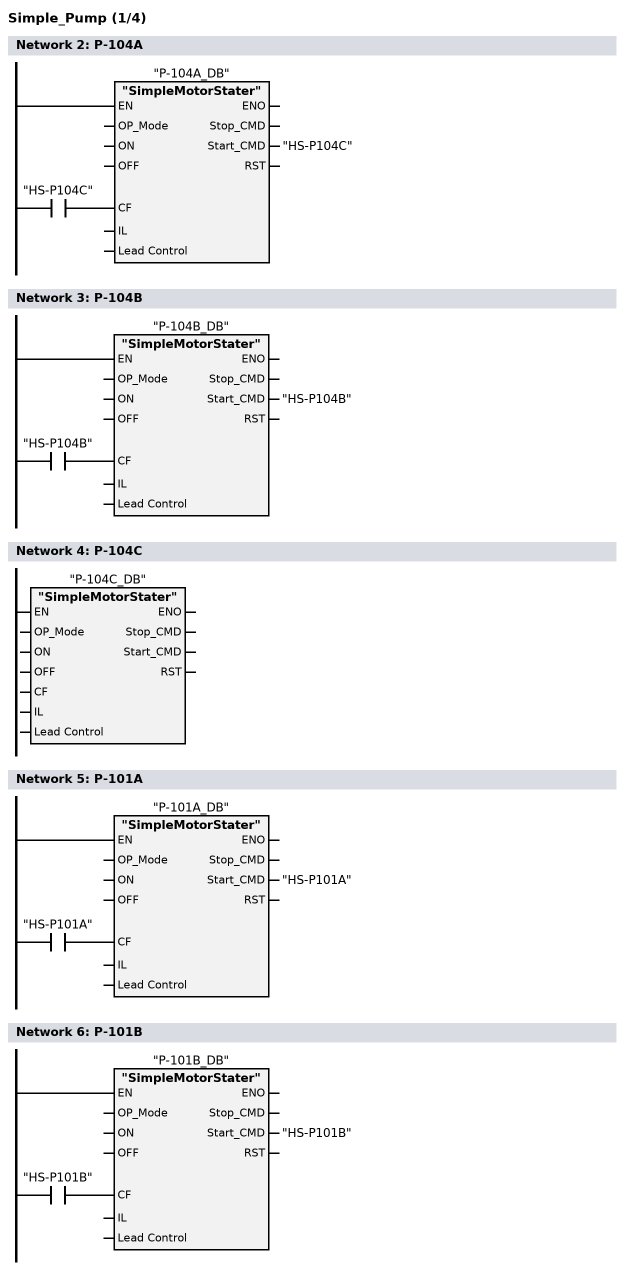
   RUNG wire#powerrail
      "P-104A_DB"(CF := wire#w1, OP_Mode :=, ON :=, OFF :=, IL :=, "Lead Control" :=, Stop_CMD =>, Start_CMD => "HS-P104C", RST =>)
   END_RUNG
   RUNG wire#powerrail
      Contact( "HS-P104C" )
   END_RUNG wire#w1
   // the same network as SCL:
   "P-104A_DB"(CF := "HS-P104C", Start_CMD => "HS-P104C");   // "SimpleMotorStater"
END_REGION

REGION Network 3: P-104B
   RUNG wire#powerrail
      "P-104B_DB"(CF := wire#w1, OP_Mode :=, ON :=, OFF :=, IL :=, "Lead Control" :=, Stop_CMD =>, Start_CMD => "HS-P104B", RST =>)
   END_RUNG
   RUNG wire#powerrail
      Contact( "HS-P104B" )
   END_RUNG wire#w1
   // the same network as SCL:
   "P-104B_DB"(CF := "HS-P104B", Start_CMD => "HS-P104B");   // "SimpleMotorStater"
END_REGION

REGION Network 4: P-104C
   RUNG wire#powerrail
      "P-104C_DB"(OP_Mode :=, ON :=, OFF :=, CF :=, IL :=, "Lead Control" :=, Stop_CMD =>, Start_CMD =>, RST =>)
   END_RUNG
   // the same network as SCL:
   "P-104C_DB"();   // "SimpleMotorStater"
END_REGION

REGION Network 5: P-101A
   RUNG wire#powerrail
      "P-101A_DB"(CF := wire#w1, OP_Mode :=, ON :=, OFF :=, IL :=, "Lead Control" :=, Stop_CMD =>, Start_CMD => "HS-P101A", RST =>)
   END_RUNG
   RUNG wire#powerrail
      Contact( "HS-P101A" )
   END_RUNG wire#w1
   // the same network as SCL:
   "P-101A_DB"(CF := "HS-P101A", Start_CMD => "HS-P101A");   // "SimpleMotorStater"
END_REGION

REGION Network 6: P-101B
   RUNG wire#powerrail
      "P-101B_DB"(CF := wire#w1, OP_Mode :=, ON :=, OFF :=, IL :=, "Lead Control" :=, Stop_CMD =>, Start_CMD => "HS-P101B", RST =>)
   END_RUNG
   RUNG wire#powerrail
      Contact( "HS-P101B" )
   END_RUNG wire#w1
   // the same network as SCL:
   "P-101B_DB"(CF := "HS-P101B", Start_CMD => "HS-P101B");   // "SimpleMotorStater"
END_REGION

REGION Network 7: P-102A
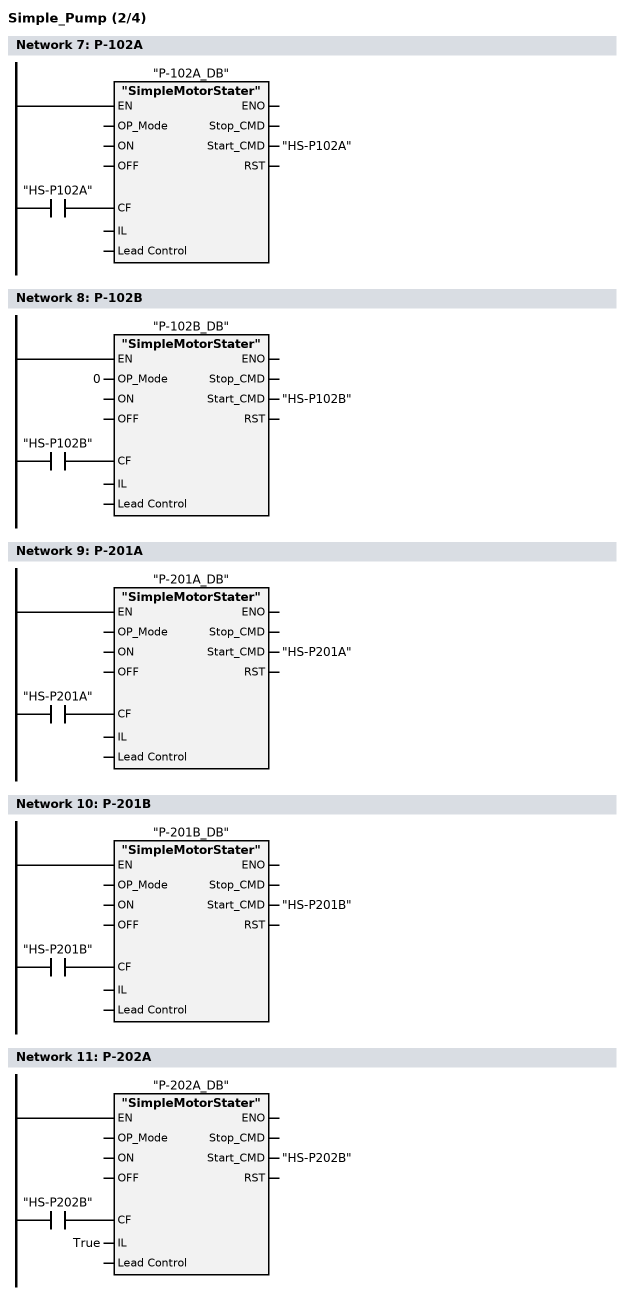
   RUNG wire#powerrail
      "P-102A_DB"(CF := wire#w1, OP_Mode :=, ON :=, OFF :=, IL :=, "Lead Control" :=, Stop_CMD =>, Start_CMD => "HS-P102A", RST =>)
   END_RUNG
   RUNG wire#powerrail
      Contact( "HS-P102A" )
   END_RUNG wire#w1
   // the same network as SCL:
   "P-102A_DB"(CF := "HS-P102A", Start_CMD => "HS-P102A");   // "SimpleMotorStater"
END_REGION

REGION Network 8: P-102B
   RUNG wire#powerrail
      "P-102B_DB"(CF := wire#w1, OP_Mode := 0, ON :=, OFF :=, IL :=, "Lead Control" :=, Stop_CMD =>, Start_CMD => "HS-P102B", RST =>)
   END_RUNG
   RUNG wire#powerrail
      Contact( "HS-P102B" )
   END_RUNG wire#w1
   // the same network as SCL:
   "P-102B_DB"(OP_Mode := 0, CF := "HS-P102B", Start_CMD => "HS-P102B");   // "SimpleMotorStater"
END_REGION

REGION Network 9: P-201A
   RUNG wire#powerrail
      "P-201A_DB"(CF := wire#w1, OP_Mode :=, ON :=, OFF :=, IL :=, "Lead Control" :=, Stop_CMD =>, Start_CMD => "HS-P201A", RST =>)
   END_RUNG
   RUNG wire#powerrail
      Contact( "HS-P201A" )
   END_RUNG wire#w1
   // the same network as SCL:
   "P-201A_DB"(CF := "HS-P201A", Start_CMD => "HS-P201A");   // "SimpleMotorStater"
END_REGION

REGION Network 10: P-201B
   RUNG wire#powerrail
      "P-201B_DB"(CF := wire#w1, OP_Mode :=, ON :=, OFF :=, IL :=, "Lead Control" :=, Stop_CMD =>, Start_CMD => "HS-P201B", RST =>)
   END_RUNG
   RUNG wire#powerrail
      Contact( "HS-P201B" )
   END_RUNG wire#w1
   // the same network as SCL:
   "P-201B_DB"(CF := "HS-P201B", Start_CMD => "HS-P201B");   // "SimpleMotorStater"
END_REGION

REGION Network 11: P-202A
   RUNG wire#powerrail
      "P-202A_DB"(CF := wire#w1, OP_Mode :=, ON :=, OFF :=, IL := True, "Lead Control" :=, Stop_CMD =>, Start_CMD => "HS-P202B", RST =>)
   END_RUNG
   RUNG wire#powerrail
      Contact( "HS-P202B" )
   END_RUNG wire#w1
   // the same network as SCL:
   "P-202A_DB"(CF := "HS-P202B", IL := True, Start_CMD => "HS-P202B");   // "SimpleMotorStater"
END_REGION

REGION Network 12: P-202B
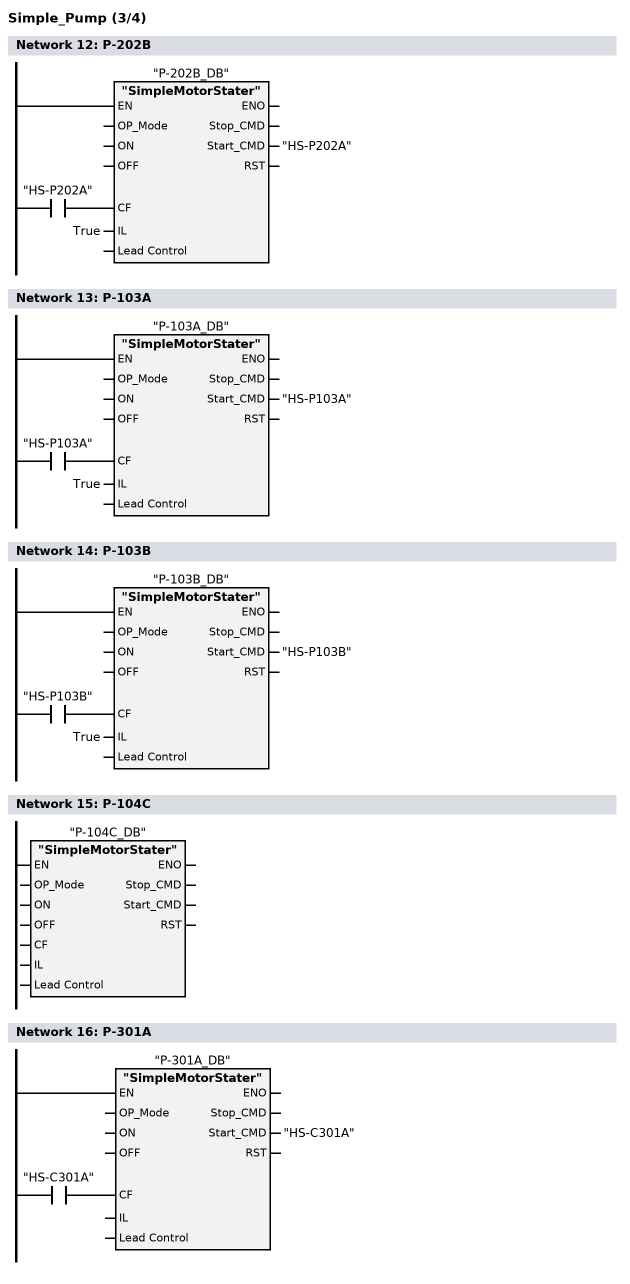
   RUNG wire#powerrail
      "P-202B_DB"(CF := wire#w1, OP_Mode :=, ON :=, OFF :=, IL := True, "Lead Control" :=, Stop_CMD =>, Start_CMD => "HS-P202A", RST =>)
   END_RUNG
   RUNG wire#powerrail
      Contact( "HS-P202A" )
   END_RUNG wire#w1
   // the same network as SCL:
   "P-202B_DB"(CF := "HS-P202A", IL := True, Start_CMD => "HS-P202A");   // "SimpleMotorStater"
END_REGION

REGION Network 13: P-103A
   RUNG wire#powerrail
      "P-103A_DB"(CF := wire#w1, OP_Mode :=, ON :=, OFF :=, IL := True, "Lead Control" :=, Stop_CMD =>, Start_CMD => "HS-P103A", RST =>)
   END_RUNG
   RUNG wire#powerrail
      Contact( "HS-P103A" )
   END_RUNG wire#w1
   // the same network as SCL:
   "P-103A_DB"(CF := "HS-P103A", IL := True, Start_CMD => "HS-P103A");   // "SimpleMotorStater"
END_REGION

REGION Network 14: P-103B
   RUNG wire#powerrail
      "P-103B_DB"(CF := wire#w1, OP_Mode :=, ON :=, OFF :=, IL := True, "Lead Control" :=, Stop_CMD =>, Start_CMD => "HS-P103B", RST =>)
   END_RUNG
   RUNG wire#powerrail
      Contact( "HS-P103B" )
   END_RUNG wire#w1
   // the same network as SCL:
   "P-103B_DB"(CF := "HS-P103B", IL := True, Start_CMD => "HS-P103B");   // "SimpleMotorStater"
END_REGION

REGION Network 15: P-104C
   RUNG wire#powerrail
      "P-104C_DB"(OP_Mode :=, ON :=, OFF :=, CF :=, IL :=, "Lead Control" :=, Stop_CMD =>, Start_CMD =>, RST =>)
   END_RUNG
   // the same network as SCL:
   "P-104C_DB"();   // "SimpleMotorStater"
END_REGION

REGION Network 16: P-301A
   RUNG wire#powerrail
      "P-301A_DB"(CF := wire#w1, OP_Mode :=, ON :=, OFF :=, IL :=, "Lead Control" :=, Stop_CMD =>, Start_CMD => "HS-C301A", RST =>)
   END_RUNG
   RUNG wire#powerrail
      Contact( "HS-C301A" )
   END_RUNG wire#w1
   // the same network as SCL:
   "P-301A_DB"(CF := "HS-C301A", Start_CMD => "HS-C301A");   // "SimpleMotorStater"
END_REGION

REGION Network 17: P-301B
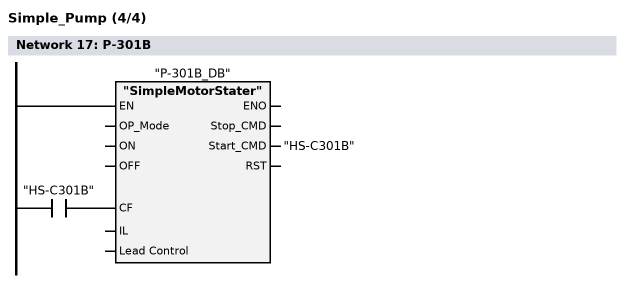
   RUNG wire#powerrail
      "P-301B_DB"(CF := wire#w1, OP_Mode :=, ON :=, OFF :=, IL :=, "Lead Control" :=, Stop_CMD =>, Start_CMD => "HS-C301B", RST =>)
   END_RUNG
   RUNG wire#powerrail
      Contact( "HS-C301B" )
   END_RUNG wire#w1
   // the same network as SCL:
   "P-301B_DB"(CF := "HS-C301B", Start_CMD => "HS-C301B");   // "SimpleMotorStater"
END_REGION
END_FUNCTION

// folder: Signal Digital Output/Centrifuge

FUNCTION "Centrifuge_DO" : Void   // FC108, LAD
{ S7_Optimized_Access := 'TRUE' }
VERSION : 0.1
BEGIN

REGION Network 1: Centrifuge Start Command
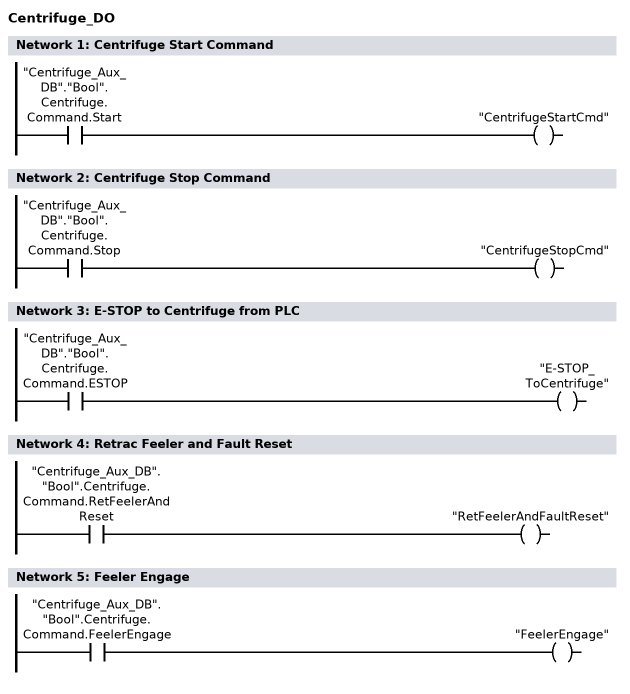
   RUNG wire#powerrail
      Contact( "Centrifuge_Aux_DB"."Bool".Centrifuge.Command.Start )
      Coil( "CentrifugeStartCmd" )
   END_RUNG
   // the same network as SCL:
   "CentrifugeStartCmd" := "Centrifuge_Aux_DB"."Bool".Centrifuge.Command.Start;
END_REGION

REGION Network 2: Centrifuge Stop Command
   RUNG wire#powerrail
      Contact( "Centrifuge_Aux_DB"."Bool".Centrifuge.Command.Stop )
      Coil( "CentrifugeStopCmd" )
   END_RUNG
   // the same network as SCL:
   "CentrifugeStopCmd" := "Centrifuge_Aux_DB"."Bool".Centrifuge.Command.Stop;
END_REGION

REGION Network 3: E-STOP to Centrifuge from PLC
   RUNG wire#powerrail
      Contact( "Centrifuge_Aux_DB"."Bool".Centrifuge.Command.ESTOP )
      Coil( "E-STOP_ToCentrifuge" )
   END_RUNG
   // the same network as SCL:
   "E-STOP_ToCentrifuge" := "Centrifuge_Aux_DB"."Bool".Centrifuge.Command.ESTOP;
END_REGION

REGION Network 4: Retrac Feeler and Fault Reset
   RUNG wire#powerrail
      Contact( "Centrifuge_Aux_DB"."Bool".Centrifuge.Command.RetFeelerAndReset )
      Coil( "RetFeelerAndFaultReset" )
   END_RUNG
   // the same network as SCL:
   "RetFeelerAndFaultReset" := "Centrifuge_Aux_DB"."Bool".Centrifuge.Command.RetFeelerAndReset;
END_REGION

REGION Network 5: Feeler Engage
   RUNG wire#powerrail
      Contact( "Centrifuge_Aux_DB"."Bool".Centrifuge.Command.FeelerEngage )
      Coil( "FeelerEngage" )
   END_RUNG
   // the same network as SCL:
   "FeelerEngage" := "Centrifuge_Aux_DB"."Bool".Centrifuge.Command.FeelerEngage;
END_REGION
END_FUNCTION

// folder: Signal Inputs

FUNCTION "Signals" : Void   // FC6, LAD
{ S7_Optimized_Access := 'TRUE' }
VERSION : 0.1
BEGIN

REGION Network 1: LSHH-1011 : T-101 High High Level Switch
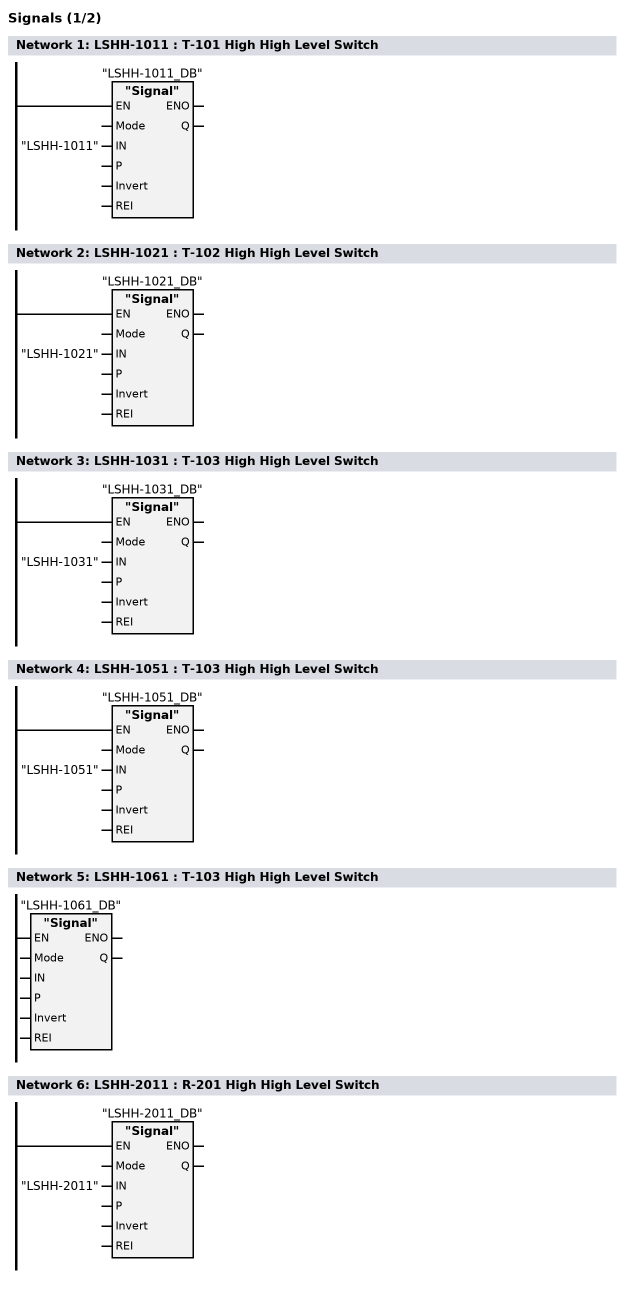
   RUNG wire#powerrail
      "LSHH-1011_DB"(Mode :=, IN := "LSHH-1011", P :=, Invert :=, REI :=, Q =>)
   END_RUNG
   // the same network as SCL:
   "LSHH-1011_DB"(IN := "LSHH-1011");   // "Signal"
END_REGION

REGION Network 2: LSHH-1021 : T-102 High High Level Switch
   RUNG wire#powerrail
      "LSHH-1021_DB"(Mode :=, IN := "LSHH-1021", P :=, Invert :=, REI :=, Q =>)
   END_RUNG
   // the same network as SCL:
   "LSHH-1021_DB"(IN := "LSHH-1021");   // "Signal"
END_REGION

REGION Network 3: LSHH-1031 : T-103 High High Level Switch
   RUNG wire#powerrail
      "LSHH-1031_DB"(Mode :=, IN := "LSHH-1031", P :=, Invert :=, REI :=, Q =>)
   END_RUNG
   // the same network as SCL:
   "LSHH-1031_DB"(IN := "LSHH-1031");   // "Signal"
END_REGION

REGION Network 4: LSHH-1051 : T-103 High High Level Switch
   RUNG wire#powerrail
      "LSHH-1051_DB"(Mode :=, IN := "LSHH-1051", P :=, Invert :=, REI :=, Q =>)
   END_RUNG
   // the same network as SCL:
   "LSHH-1051_DB"(IN := "LSHH-1051");   // "Signal"
END_REGION

REGION Network 5: LSHH-1061 : T-103 High High Level Switch
   RUNG wire#powerrail
      "LSHH-1061_DB"(Mode :=, IN :=, P :=, Invert :=, REI :=, Q =>)
   END_RUNG
   // the same network as SCL:
   "LSHH-1061_DB"();   // "Signal"
END_REGION

REGION Network 6: LSHH-2011 : R-201 High High Level Switch
   RUNG wire#powerrail
      "LSHH-2011_DB"(Mode :=, IN := "LSHH-2011", P :=, Invert :=, REI :=, Q =>)
   END_RUNG
   // the same network as SCL:
   "LSHH-2011_DB"(IN := "LSHH-2011");   // "Signal"
END_REGION

REGION Network 7: LSHH-2021 : R-202 High High Level Switch
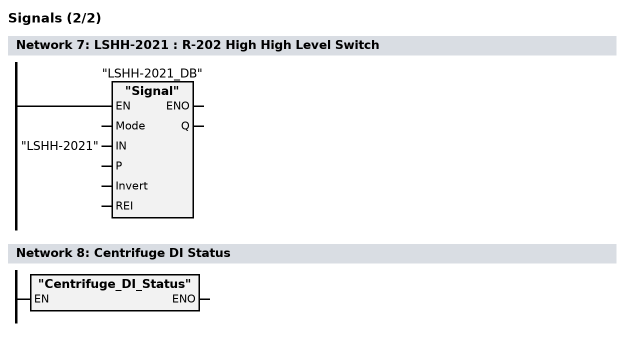
   RUNG wire#powerrail
      "LSHH-2021_DB"(Mode :=, IN := "LSHH-2021", P :=, Invert :=, REI :=, Q =>)
   END_RUNG
   // the same network as SCL:
   "LSHH-2021_DB"(IN := "LSHH-2021");   // "Signal"
END_REGION

REGION Network 8: Centrifuge DI Status
   RUNG wire#powerrail
      "Centrifuge_DI_Status"()
   END_RUNG
   // the same network as SCL:
   "Centrifuge_DI_Status"();
END_REGION
END_FUNCTION

// folder: Signal Inputs/Centrifuge

FUNCTION "Centrifuge_DI_Status" : Void   // FC104, LAD
{ S7_Optimized_Access := 'TRUE' }
VERSION : 0.1
// Digital Input from Centrifuge
BEGIN

REGION Network 1: Vibration Fault
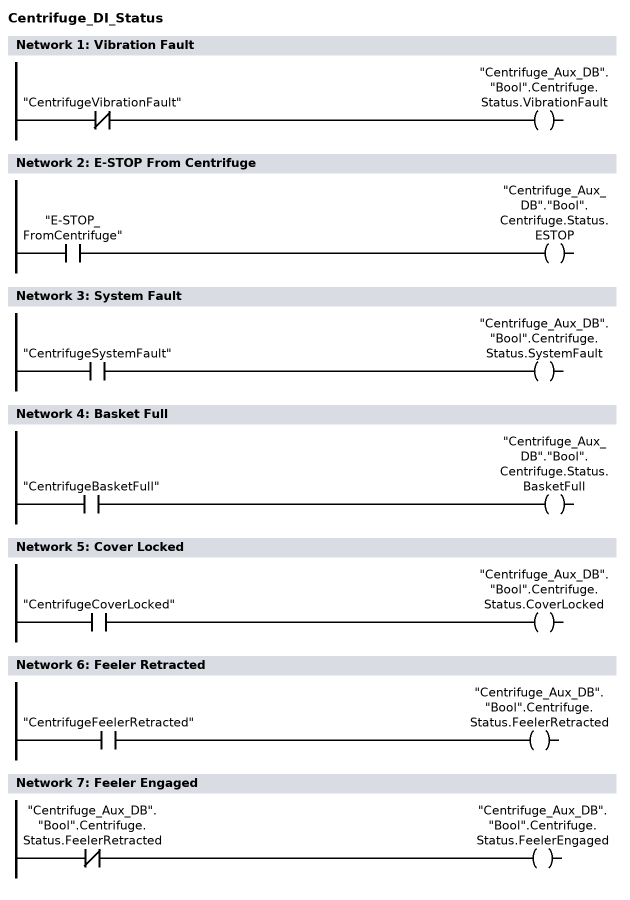
   RUNG wire#powerrail
      I_Contact( "CentrifugeVibrationFault" )
      Coil( "Centrifuge_Aux_DB"."Bool".Centrifuge.Status.VibrationFault )
   END_RUNG
   // the same network as SCL:
   "Centrifuge_Aux_DB"."Bool".Centrifuge.Status.VibrationFault := NOT "CentrifugeVibrationFault";
END_REGION

REGION Network 2: E-STOP From Centrifuge
   RUNG wire#powerrail
      Contact( "E-STOP_FromCentrifuge" )
      Coil( "Centrifuge_Aux_DB"."Bool".Centrifuge.Status.ESTOP )
   END_RUNG
   // the same network as SCL:
   "Centrifuge_Aux_DB"."Bool".Centrifuge.Status.ESTOP := "E-STOP_FromCentrifuge";
END_REGION

REGION Network 3: System Fault
   RUNG wire#powerrail
      Contact( "CentrifugeSystemFault" )
      Coil( "Centrifuge_Aux_DB"."Bool".Centrifuge.Status.SystemFault )
   END_RUNG
   // the same network as SCL:
   "Centrifuge_Aux_DB"."Bool".Centrifuge.Status.SystemFault := "CentrifugeSystemFault";
END_REGION

REGION Network 4: Basket Full
   RUNG wire#powerrail
      Contact( "CentrifugeBasketFull" )
      Coil( "Centrifuge_Aux_DB"."Bool".Centrifuge.Status.BasketFull )
   END_RUNG
   // the same network as SCL:
   "Centrifuge_Aux_DB"."Bool".Centrifuge.Status.BasketFull := "CentrifugeBasketFull";
END_REGION

REGION Network 5: Cover Locked
   RUNG wire#powerrail
      Contact( "CentrifugeCoverLocked" )
      Coil( "Centrifuge_Aux_DB"."Bool".Centrifuge.Status.CoverLocked )
   END_RUNG
   // the same network as SCL:
   "Centrifuge_Aux_DB"."Bool".Centrifuge.Status.CoverLocked := "CentrifugeCoverLocked";
END_REGION

REGION Network 6: Feeler Retracted
   RUNG wire#powerrail
      Contact( "CentrifugeFeelerRetracted" )
      Coil( "Centrifuge_Aux_DB"."Bool".Centrifuge.Status.FeelerRetracted )
   END_RUNG
   // the same network as SCL:
   "Centrifuge_Aux_DB"."Bool".Centrifuge.Status.FeelerRetracted := "CentrifugeFeelerRetracted";
END_REGION

REGION Network 7: Feeler Engaged
   RUNG wire#powerrail
      I_Contact( "Centrifuge_Aux_DB"."Bool".Centrifuge.Status.FeelerRetracted )
      Coil( "Centrifuge_Aux_DB"."Bool".Centrifuge.Status.FeelerEngaged )
   END_RUNG
   // the same network as SCL:
   "Centrifuge_Aux_DB"."Bool".Centrifuge.Status.FeelerEngaged := NOT "Centrifuge_Aux_DB"."Bool".Centrifuge.Status.FeelerRetracted;
END_REGION
END_FUNCTION

// folder: State MACHINE

FUNCTION "Sequence_Caller" : Void   // FC39, LAD
{ S7_Optimized_Access := 'TRUE' }
VERSION : 0.1
BEGIN

REGION Network 1: R-201 Reactor Control SEQ
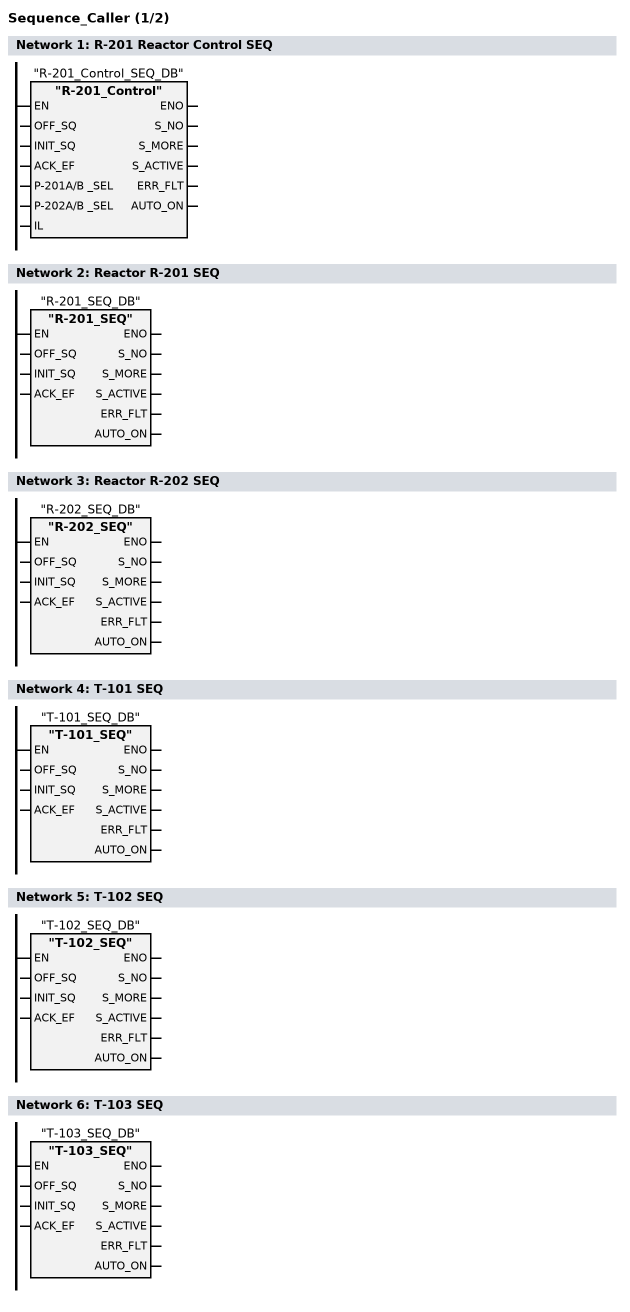
   RUNG wire#powerrail
      "R-201_Control_SEQ_DB"(OFF_SQ :=, INIT_SQ :=, ACK_EF :=, "P-201A/B _SEL" :=, "P-202A/B _SEL" :=, IL :=, S_NO =>, S_MORE =>, S_ACTIVE =>, ERR_FLT =>, AUTO_ON =>)
   END_RUNG
   // the same network as SCL:
   "R-201_Control_SEQ_DB"();   // "R-201_Control"
END_REGION

REGION Network 2: Reactor R-201 SEQ
   RUNG wire#powerrail
      "R-201_SEQ_DB"(OFF_SQ :=, INIT_SQ :=, ACK_EF :=, S_NO =>, S_MORE =>, S_ACTIVE =>, ERR_FLT =>, AUTO_ON =>)
   END_RUNG
   // the same network as SCL:
   "R-201_SEQ_DB"();   // "R-201_SEQ"
END_REGION

REGION Network 3: Reactor R-202 SEQ
   RUNG wire#powerrail
      "R-202_SEQ_DB"(OFF_SQ :=, INIT_SQ :=, ACK_EF :=, S_NO =>, S_MORE =>, S_ACTIVE =>, ERR_FLT =>, AUTO_ON =>)
   END_RUNG
   // the same network as SCL:
   "R-202_SEQ_DB"();   // "R-202_SEQ"
END_REGION

REGION Network 4: T-101 SEQ
   RUNG wire#powerrail
      "T-101_SEQ_DB"(OFF_SQ :=, INIT_SQ :=, ACK_EF :=, S_NO =>, S_MORE =>, S_ACTIVE =>, ERR_FLT =>, AUTO_ON =>)
   END_RUNG
   // the same network as SCL:
   "T-101_SEQ_DB"();   // "T-101_SEQ"
END_REGION

REGION Network 5: T-102 SEQ
   RUNG wire#powerrail
      "T-102_SEQ_DB"(OFF_SQ :=, INIT_SQ :=, ACK_EF :=, S_NO =>, S_MORE =>, S_ACTIVE =>, ERR_FLT =>, AUTO_ON =>)
   END_RUNG
   // the same network as SCL:
   "T-102_SEQ_DB"();   // "T-102_SEQ"
END_REGION

REGION Network 6: T-103 SEQ
   RUNG wire#powerrail
      "T-103_SEQ_DB"(OFF_SQ :=, INIT_SQ :=, ACK_EF :=, S_NO =>, S_MORE =>, S_ACTIVE =>, ERR_FLT =>, AUTO_ON =>)
   END_RUNG
   // the same network as SCL:
   "T-103_SEQ_DB"();   // "T-103_SEQ"
END_REGION

REGION Network 7: T-104 SEQ
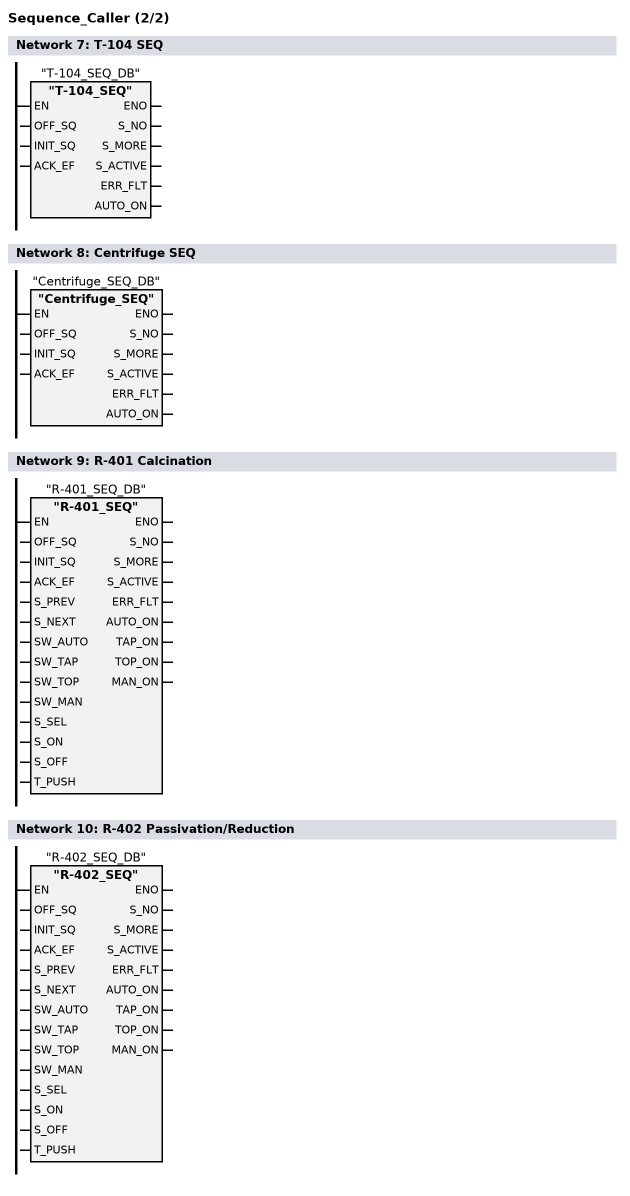
   RUNG wire#powerrail
      "T-104_SEQ_DB"(OFF_SQ :=, INIT_SQ :=, ACK_EF :=, S_NO =>, S_MORE =>, S_ACTIVE =>, ERR_FLT =>, AUTO_ON =>)
   END_RUNG
   // the same network as SCL:
   "T-104_SEQ_DB"();   // "T-104_SEQ"
END_REGION

REGION Network 8: Centrifuge SEQ
   RUNG wire#powerrail
      "Centrifuge_SEQ_DB"(OFF_SQ :=, INIT_SQ :=, ACK_EF :=, S_NO =>, S_MORE =>, S_ACTIVE =>, ERR_FLT =>, AUTO_ON =>)
   END_RUNG
   // the same network as SCL:
   "Centrifuge_SEQ_DB"();   // "Centrifuge_SEQ"
END_REGION

REGION Network 9: R-401 Calcination
   RUNG wire#powerrail
      "R-401_SEQ_DB"(OFF_SQ :=, INIT_SQ :=, ACK_EF :=, S_PREV :=, S_NEXT :=, SW_AUTO :=, SW_TAP :=, SW_TOP :=, SW_MAN :=, S_SEL :=, S_ON :=, S_OFF :=, T_PUSH :=, S_NO =>, S_MORE =>, S_ACTIVE =>, ERR_FLT =>, AUTO_ON =>, TAP_ON =>, TOP_ON =>, MAN_ON =>)
   END_RUNG
   // the same network as SCL:
   "R-401_SEQ_DB"();   // "R-401_SEQ"
END_REGION

REGION Network 10: R-402 Passivation/Reduction
   RUNG wire#powerrail
      "R-402_SEQ_DB"(OFF_SQ :=, INIT_SQ :=, ACK_EF :=, S_PREV :=, S_NEXT :=, SW_AUTO :=, SW_TAP :=, SW_TOP :=, SW_MAN :=, S_SEL :=, S_ON :=, S_OFF :=, T_PUSH :=, S_NO =>, S_MORE =>, S_ACTIVE =>, ERR_FLT =>, AUTO_ON =>, TAP_ON =>, TOP_ON =>, MAN_ON =>)
   END_RUNG
   // the same network as SCL:
   "R-402_SEQ_DB"();   // "R-402_SEQ"
END_REGION
END_FUNCTION

// folder: State MACHINE/1)Tanks/Tank T-101 (X)

FUNCTION_BLOCK "T-101_SEQ"   // FB41, GRAPH_PLUS
{ S7_Optimized_Access := 'TRUE' }
VERSION : 0.1
   VAR_INPUT
      OFF_SQ : Bool := false;   // Turn sequence off
      INIT_SQ : Bool := false;   // Set sequence to initial state
      ACK_EF : Bool := false;   // Acknowledge all errors and faults
   END_VAR
   VAR_OUTPUT
      S_NO : Int := 0;   // Step number
      S_MORE : Bool := false;   // More steps are available and can be shown in S_NO
      S_ACTIVE : Bool := false;   // Step indicated in S_NO is active
      ERR_FLT : Bool := false;   // Interlock or supervision group error
      AUTO_ON : Bool := false;   // Automatic mode is active
   END_VAR
   VAR
      HMI_INFO : Array[0..10] of UInt;
      IF_PAR : G7_IfParPlus_V6;
      RT_DATA : G7_RTDataPlus_V6;   // Internal data area
      Abort : G7_TransitionPlus_V6;   // Transition structure
      InitializeTk : G7_TransitionPlus_V6;   // Transition structure
      Block : G7_TransitionPlus_V6;   // Transition structure
      Rdy : G7_TransitionPlus_V6;   // Transition structure
      MixSeq : G7_TransitionPlus_V6;   // Transition structure
      WashSeq : G7_TransitionPlus_V6;   // Transition structure
      Pouring : G7_TransitionPlus_V6;   // Transition structure
      Started : G7_TransitionPlus_V6;   // Transition structure
      Params : G7_TransitionPlus_V6;   // Transition structure
      FillingDn : G7_TransitionPlus_V6;   // Transition structure
      WaterOff : G7_TransitionPlus_V6;   // Transition structure
      TankR : G7_TransitionPlus_V6;   // Transition structure
      "Open Signal_1" : G7_TransitionPlus_V6;   // Transition structure
      MixTimeDn : G7_TransitionPlus_V6;   // Transition structure
      MixOpDn : G7_TransitionPlus_V6;   // Transition structure
      NoFlow : G7_TransitionPlus_V6;   // Transition structure
      MixDn : G7_TransitionPlus_V6;   // Transition structure
      PourSt : G7_TransitionPlus_V6;   // Transition structure
      Rc : G7_TransitionPlus_V6;   // Transition structure
      Transf : G7_TransitionPlus_V6;   // Transition structure
      ClsR : G7_TransitionPlus_V6;   // Transition structure
      Release : G7_TransitionPlus_V6;   // Transition structure
      Init : G7_TransitionPlus_V6;   // Transition structure
      SAut : G7_TransitionPlus_V6;   // Transition structure
      SIn : G7_TransitionPlus_V6;   // Transition structure
      Initd : G7_TransitionPlus_V6;   // Transition structure
      Ab : G7_TransitionPlus_V6;   // Transition structure
      AbortOn : G7_TransitionPlus_V6;   // Transition structure
      AbortDn : G7_TransitionPlus_V6;   // Transition structure
      Idle : G7_StepPlus_V6;   // Step structure
      Ready : G7_StepPlus_V6;   // Step structure
      SelectSeq : G7_StepPlus_V6;   // Step structure
      MixStarted : G7_StepPlus_V6;   // Step structure
      "EDIT QWater" : G7_StepPlus_V6;   // Step structure
      FillingUpWater : G7_StepPlus_V6;   // Step structure
      StopReqWater : G7_StepPlus_V6;   // Step structure
      "ReleaseT-104" : G7_StepPlus_V6;   // Step structure
      "USER PourDn" : G7_StepPlus_V6;   // Step structure
      MinMixingTime : G7_StepPlus_V6;   // Step structure
      "USER EndMix" : G7_StepPlus_V6;   // Step structure
      ShuttingDown : G7_StepPlus_V6;   // Step structure
      DoneMix : G7_StepPlus_V6;   // Step structure
      PouringStarted : G7_StepPlus_V6;   // Step structure
      Recirculation : G7_StepPlus_V6;   // Step structure
      Transfering : G7_StepPlus_V6;   // Step structure
      CloseRoute : G7_StepPlus_V6;   // Step structure
      DoneTransfer : G7_StepPlus_V6;   // Step structure
      Initialize : G7_StepPlus_V6;   // Step structure
      SetAuto : G7_StepPlus_V6;   // Step structure
      SetInitial : G7_StepPlus_V6;   // Step structure
      Initialized : G7_StepPlus_V6;   // Step structure
      AbortStarting : G7_StepPlus_V6;   // Step structure
      Aborting : G7_StepPlus_V6;   // Step structure
      Abort_Done : G7_StepPlus_V6;   // Step structure
      SINI : Array[0..3] of USInt;
      LSTT : Array[0..28] of USInt;
      ATAJ : Array[0..28] of USInt;
      ATAB : Array[0..28] of USInt;
      PSTT : Array[0..28] of USInt;
      NSTT : Array[0..28] of USInt;
      ASSJ : Array[0..24] of USInt;
      ASSB : Array[0..24] of USInt;
      PTTS : Array[0..24] of USInt;
      NTTS : Array[0..24] of USInt;
      SW_SQTS : Array[0..24] of USInt;
      SWITCH : Array[0..4] of USInt;
      TVX : Array[0..9] of USInt;
      TTX : Array[0..9] of USInt;
      TSX : Array[0..3] of USInt;
      S00X : Array[0..3] of USInt;
      SOFFX : Array[0..3] of USInt;
      SONX : Array[0..3] of USInt;
      SAX : Array[0..3] of USInt;
      SERRX : Array[0..25] of USInt;
      SMX : Array[0..25] of USInt;
      S0X : Array[0..25] of USInt;
      S1X : Array[0..25] of USInt;
      IL_ALARM_INST : Diag_Alarm;
      SUP_ALARM_INST : Diag_Alarm;
      STEP_TIME_ALARM_INST : Diag_Alarm;
      IEC_TIMER_INST : IEC_TIMER;
      TRANSACTION_FLAG : Bool := false;
   END_VAR
   // SINI[0] := 2;
   // SINI[2] := 255;
   // SINI[3] := 255;
   // LSTT[0] := 22;
   // LSTT[1] := 18;
   // LSTT[2] := 255;
   // LSTT[3] := 255;
   // LSTT[4] := 255;
   // LSTT[12] := 255;
   // LSTT[6] := 255;
   // LSTT[7] := 255;
   // LSTT[8] := 255;
   // LSTT[9] := 255;
   // LSTT[10] := 255;
   // LSTT[11] := 255;
   // LSTT[13] := 255;
   // LSTT[15] := 255;
   // LSTT[20] := 255;
   // LSTT[17] := 255;
   // LSTT[18] := 255;
   // LSTT[19] := 255;
   // LSTT[27] := 255;
   // LSTT[22] := 255;
   // LSTT[23] := 255;
   // LSTT[24] := 255;
   // LSTT[25] := 1;
   // LSTT[26] := 255;
   // NSTT[14] := 11;
   // ATAJ[1] := 1;
   // ATAJ[2] := 2;
   // ATAJ[3] := 3;
   // ATAJ[4] := 4;
   // ATAJ[5] := 5;
   // ATAJ[6] := 6;
   // ATAJ[7] := 7;
   // ATAJ[8] := 8;
   // ATAJ[9] := 9;
   // ATAJ[10] := 10;
   // ATAJ[11] := 11;
   // ATAJ[12] := 12;
   // ATAJ[13] := 13;
   // ATAJ[14] := 14;
   // ATAJ[15] := 15;
   // ATAJ[16] := 16;
   // ATAJ[17] := 17;
   // ATAJ[18] := 18;
   // ATAJ[19] := 19;
   // ATAJ[20] := 20;
   // ATAJ[21] := 21;
   // ATAJ[22] := 22;
   // ATAJ[23] := 23;
   // ATAJ[24] := 24;
   // ATAJ[25] := 25;
   // ATAJ[26] := 26;
   // ATAJ[27] := 27;
   // ATAJ[28] := 28;
   // ATAB[0] := 1;
   // ATAB[1] := 2;
   // ATAB[24] := 24;
   // ATAB[3] := 3;
   // ATAB[4] := 5;
   // ATAB[5] := 6;
   // ATAB[6] := 4;
   // ATAB[7] := 7;
   // ATAB[8] := 8;
   // ATAB[9] := 9;
   // ATAB[10] := 10;
   // ATAB[11] := 11;
   // ATAB[12] := 12;
   // ATAB[13] := 13;
   // ATAB[14] := 14;
   // ATAB[15] := 15;
   // ATAB[16] := 16;
   // ATAB[17] := 17;
   // ATAB[18] := 18;
   // ATAB[19] := 19;
   // ATAB[20] := 20;
   // ATAB[21] := 21;
   // ATAB[22] := 22;
   // ATAB[23] := 23;
   // ATAB[25] := 25;
   // ATAB[26] := 26;
   // ATAB[27] := 27;
   // ATAB[28] := 28;
   // PSTT[24] := 20;
   // PSTT[5] := 2;
   // PSTT[3] := 1;
   // PSTT[4] := 2;
   // PSTT[15] := 11;
   // PSTT[6] := 2;
   // PSTT[7] := 3;
   // PSTT[8] := 4;
   // PSTT[9] := 5;
   // PSTT[10] := 6;
   // PSTT[11] := 7;
   // PSTT[12] := 8;
   // PSTT[13] := 9;
   // PSTT[14] := 10;
   // PSTT[16] := 12;
   // PSTT[17] := 13;
   // PSTT[18] := 14;
   // PSTT[19] := 15;
   // PSTT[20] := 16;
   // PSTT[21] := 17;
   // PSTT[22] := 18;
   // PSTT[23] := 19;
   // PSTT[25] := 21;
   // PSTT[26] := 22;
   // PSTT[27] := 23;
   // PSTT[28] := 24;
   // NSTT[0] := 22;
   // NSTT[1] := 18;
   // NSTT[2] := 1;
   // NSTT[3] := 2;
   // NSTT[4] := 3;
   // NSTT[12] := 9;
   // NSTT[6] := 13;
   // NSTT[7] := 4;
   // NSTT[8] := 5;
   // NSTT[9] := 6;
   // NSTT[10] := 7;
   // NSTT[11] := 8;
   // NSTT[13] := 10;
   // NSTT[15] := 12;
   // NSTT[20] := 17;
   // NSTT[17] := 14;
   // NSTT[18] := 15;
   // NSTT[19] := 16;
   // NSTT[27] := 24;
   // NSTT[22] := 19;
   // NSTT[23] := 20;
   // NSTT[24] := 21;
   // NSTT[25] := 1;
   // NSTT[26] := 23;
   // ASSJ[1] := 1;
   // ASSJ[2] := 2;
   // ASSJ[3] := 3;
   // ASSJ[4] := 4;
   // ASSJ[5] := 5;
   // ASSJ[6] := 6;
   // ASSJ[7] := 7;
   // ASSJ[8] := 8;
   // ASSJ[9] := 9;
   // ASSJ[10] := 10;
   // ASSJ[11] := 11;
   // ASSJ[12] := 12;
   // ASSJ[13] := 13;
   // ASSJ[14] := 14;
   // ASSJ[15] := 15;
   // ASSJ[16] := 16;
   // ASSJ[17] := 17;
   // ASSJ[18] := 18;
   // ASSJ[19] := 19;
   // ASSJ[20] := 20;
   // ASSJ[21] := 21;
   // ASSJ[22] := 22;
   // ASSJ[23] := 23;
   // ASSJ[24] := 24;
   // ASSB[1] := 1;
   // ASSB[2] := 2;
   // ASSB[3] := 3;
   // ASSB[4] := 4;
   // ASSB[5] := 5;
   // ASSB[6] := 6;
   // ASSB[7] := 7;
   // ASSB[8] := 8;
   // ASSB[9] := 9;
   // ASSB[10] := 10;
   // ASSB[11] := 11;
   // ASSB[12] := 12;
   // ASSB[13] := 13;
   // ASSB[14] := 14;
   // ASSB[15] := 15;
   // ASSB[16] := 16;
   // ASSB[17] := 17;
   // ASSB[18] := 18;
   // ASSB[19] := 19;
   // ASSB[20] := 20;
   // ASSB[21] := 21;
   // ASSB[22] := 22;
   // ASSB[23] := 23;
   // ASSB[24] := 24;
   // PTTS[0] := 255;
   // PTTS[1] := 2;
   // PTTS[2] := 3;
   // PTTS[3] := 4;
   // PTTS[4] := 7;
   // PTTS[5] := 8;
   // PTTS[6] := 9;
   // PTTS[7] := 10;
   // PTTS[8] := 11;
   // PTTS[9] := 12;
   // PTTS[10] := 13;
   // PTTS[11] := 14;
   // PTTS[12] := 15;
   // PTTS[13] := 6;
   // PTTS[14] := 17;
   // PTTS[15] := 18;
   // PTTS[16] := 19;
   // PTTS[17] := 20;
   // PTTS[18] := 255;
   // PTTS[19] := 22;
   // PTTS[20] := 23;
   // PTTS[21] := 24;
   // PTTS[22] := 255;
   // PTTS[23] := 26;
   // PTTS[24] := 27;
   // NTTS[1] := 3;
   // NTTS[2] := 4;
   // NTTS[3] := 7;
   // NTTS[4] := 8;
   // NTTS[5] := 9;
   // NTTS[6] := 10;
   // NTTS[7] := 11;
   // NTTS[8] := 12;
   // NTTS[9] := 13;
   // NTTS[10] := 14;
   // NTTS[11] := 15;
   // NTTS[12] := 16;
   // NTTS[13] := 17;
   // NTTS[14] := 18;
   // NTTS[15] := 19;
   // NTTS[16] := 20;
   // NTTS[17] := 21;
   // NTTS[18] := 22;
   // NTTS[19] := 23;
   // NTTS[20] := 24;
   // NTTS[21] := 25;
   // NTTS[22] := 26;
   // NTTS[23] := 27;
   // NTTS[24] := 28;
   // SW_SQTS[1] := 1;
   // SW_SQTS[2] := 1;
   // SW_SQTS[3] := 2;
   // SW_SQTS[4] := 2;
   // SW_SQTS[5] := 2;
   // SW_SQTS[6] := 2;
   // SW_SQTS[7] := 2;
   // SW_SQTS[8] := 2;
   // SW_SQTS[9] := 2;
   // SW_SQTS[10] := 2;
   // SW_SQTS[11] := 2;
   // SW_SQTS[12] := 2;
   // SW_SQTS[13] := 3;
   // SW_SQTS[14] := 3;
   // SW_SQTS[15] := 3;
   // SW_SQTS[16] := 3;
   // SW_SQTS[17] := 3;
   // SW_SQTS[18] := 4;
   // SW_SQTS[19] := 4;
   // SW_SQTS[20] := 4;
   // SW_SQTS[21] := 4;
   // SW_SQTS[22] := 5;
   // SW_SQTS[23] := 5;
   // SW_SQTS[24] := 5;
   // SWITCH[0] := 48;
   // SWITCH[1] := 12;
   // SWITCH[2] := 195;
   // SWITCH[3] := 239;
   // SWITCH[4] := 7;
   // TVX[0] := 16#1;
   // TTX[0] := 16#1;
   // TSX[0] := 16#1;
   // S00X[0] := 16#1;
   // SOFFX[0] := 16#1;
   // SONX[0] := 16#1;
   // SAX[0] := 16#1;
   // SERRX[0] := 16#1;
   // SMX[0] := 16#1;
   // S0X[0] := 16#1;
   // S1X[0] := 16#1;
   // LSTT[14] := 255;
BEGIN
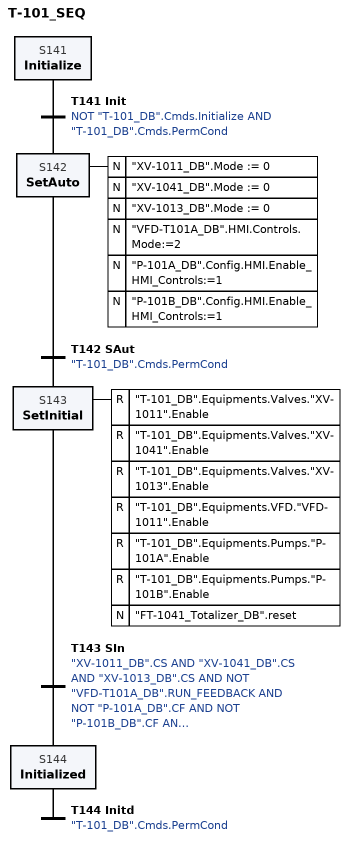
   // permanent pre-instructions
   NETWORK 1
      "T-101_Signals_FROM_R-201"();
      "T-101_Signals_FROM_R-202"();
      "T-101_Signals_FROM_T-104"();
      "T-101_SEQ_FC"();

   // sequencer 1
   STEP Initialize:   // S141, max time T#10S, warning time T#7S
      // Initialize T-101 Batch sequence
   END_STEP
   TRANSITION Init FROM Initialize TO SetAuto   // T141
      := NOT "T-101_DB".Cmds.Initialize AND "T-101_DB".Cmds.PermCond;
   END_TRANSITION
   STEP SetAuto:   // S142, max time T#10S, warning time T#7S
              N    "XV-1011_DB".Mode := 0
              N    "XV-1041_DB".Mode := 0
              N    "XV-1013_DB".Mode := 0
              N    "VFD-T101A_DB".HMI.Controls.Mode:=2
              N    "P-101A_DB".Config.HMI.Enable_HMI_Controls:=1
              N    "P-101B_DB".Config.HMI.Enable_HMI_Controls:=1
   END_STEP
   TRANSITION SAut FROM SetAuto TO SetInitial   // T142
      := "T-101_DB".Cmds.PermCond;
   END_TRANSITION
   STEP SetInitial:   // S143, max time T#10S, warning time T#7S
              R    "T-101_DB".Equipments.Valves."XV-1011".Enable
              R    "T-101_DB".Equipments.Valves."XV-1041".Enable
              R    "T-101_DB".Equipments.Valves."XV-1013".Enable
              R    "T-101_DB".Equipments.VFD."VFD-1011".Enable
              R    "T-101_DB".Equipments.Pumps."P-101A".Enable
              R    "T-101_DB".Equipments.Pumps."P-101B".Enable
              N    "FT-1041_Totalizer_DB".reset
   END_STEP
   TRANSITION SIn FROM SetInitial TO Initialized   // T143
      := "XV-1011_DB".CS AND "XV-1041_DB".CS AND "XV-1013_DB".CS AND NOT "VFD-T101A_DB".RUN_FEEDBACK AND NOT "P-101A_DB".CF AND NOT "P-101B_DB".CF AND ("FT-1041_Totalizer_DB".Total = 0.0) AND "T-101_DB".Cmds.PermCond;
   END_TRANSITION
   STEP Initialized:   // S144, max time T#10S, warning time T#7S
   END_STEP
   TRANSITION Initd FROM Initialized TO ?   // T144
      := "T-101_DB".Cmds.PermCond;
   END_TRANSITION

   // permanent post-instructions
   NETWORK 1
      "T-101_FC_Outputs"();
END_FUNCTION_BLOCK

FUNCTION "T-101_SEQ_FC" : Void   // FC53, LAD
{ S7_Optimized_Access := 'TRUE' }
VERSION : 0.1
   VAR_TEMP   // added for the SCL form of the ladder/FBD networks
      _w1 : Bool;
      _w2 : Bool;
      _w3 : Bool;
   END_VAR
BEGIN

REGION Network 2: Abort
